VERSION : 0.1
   VAR_INPUT
      SetGroup : Bool;
      "Max Seq Time h_real" : Real;
      "Max Seq Time h" : Time;
      "De-Ox Time h_real" : Real;
      "Re-Ox Time h_real" : Real;
      "Sequence Time h" : Time;
      "Setpoint Time h_real" : Real;
      "Setpoint Time h" : Time;
      "Sequence Time m Offset_real" : Real := 13.0;
      "Sequence Time m Offset" : Time;
      "O2 Confirmed Time_real" : Real;
      "O2 Confirmed Time" : Time;
      "O2 De-Ox Setpoint" : Real;
      "Re-Ox Treatment" : Bool;
      Continue : Bool;   // Continue Sequence After Restart
      Boost : Bool;   // Bypass Sequence Timers
      "Alarm Debounce time" : Time := T#30s;
      "Valve Cycle" : Struct
         Enable : Bool := true;
         Period : Time := T#2h;
         Length : Time := T#30s;
      END_STRUCT;
      "RIO 1" : "3T_IP_DATA";
      "RIO 2" : "2T_IP_DATA";
      "RIO 3" : "2T_IP_DATA";
      "RIO 4" : "2T_IP_DATA";
      "RIO 5" : "2T_IP_DATA";
      "RIO 6" : "2T_IP_DATA";
      "RIO 7" : "1T_IP_DATA";
      RUN : Bool;
      "RUN GROUP 1" : Bool;
      "RUN GROUP 2" : Bool;
      "RUN GROUP 3" : Bool;
      "RUN GROUP 4" : Bool;
      "RUN GROUP 5" : Bool;
      "RUN GROUP 6" : Bool;
      "RUN GROUP 7" : Bool;
      "RUN GROUP 8" : Bool;
      "RUN GROUP 9" : Bool;
      "RUN GROUP 10" : Bool;
      "RUN GROUP 11" : Bool;
      "RUN GROUP 12" : Bool;
      "RUN GROUP 13" : Bool;
      "RUN GROUP 14" : Bool;
      "GROUP ACTIV 1" : Bool;
      "GROUP ACTIV 2" : Bool;
      "GROUP ACTIV 3" : Bool;
      "GROUP ACTIV 4" : Bool;
      "GROUP ACTIV 5" : Bool;
      "GROUP ACTIV 6" : Bool;
      "GROUP ACTIV 7" : Bool;
      "GROUP ACTIV 8" : Bool;
      "GROUP ACTIV 9" : Bool;
      "GROUP ACTIV 10" : Bool;
      "GROUP ACTIV 11" : Bool;
      "GROUP ACTIV 12" : Bool;
      "GROUP ACTIV 13" : Bool;
      "GROUP ACTIV 14" : Bool;
      "TANK ACTIV 1" : Bool;
      "TANK ACTIV 2" : Bool;
      "TANK ACTIV 3" : Bool;
      "TANK ACTIV 4" : Bool;
      "TANK ACTIV 5" : Bool;
      "TANK ACTIV 6" : Bool;
      "TANK ACTIV 7" : Bool;
      "TANK ACTIV 8" : Bool;
      "TANK ACTIV 9" : Bool;
      "TANK ACTIV 10" : Bool;
      "TANK ACTIV 11" : Bool;
      "TANK ACTIV 12" : Bool;
      "TANK ACTIV 13" : Bool;
      "TANK ACTIV 14" : Bool;
      "TANK ACTIV 15" : Bool;
      "TANK ACTIV 16" : Bool;
      "TANK ACTIV 17" : Bool;
      "TANK ACTIV 18" : Bool;
      "TANK ACTIV 19" : Bool;
      "TANK ACTIV 20" : Bool;
      "TANK ACTIV 21" : Bool;
      "TANK ACTIV 22" : Bool;
      "TANK ACTIV 23" : Bool;
      "TANK ACTIV 24" : Bool;
   END_VAR
   VAR_OUTPUT
      "RUN TANK 1" : Bool;
      "RUN TANK 2" : Bool;
      "RUN TANK 3" : Bool;
      "RUN TANK 4" : Bool;
      "RUN TANK 5" : Bool;
      "RUN TANK 6" : Bool;
      "RUN TANK 7" : Bool;
      "RUN TANK 8" : Bool;
      "RUN TANK 9" : Bool;
      "RUN TANK 10" : Bool;
      "RUN TANK 11" : Bool;
      "RUN TANK 12" : Bool;
      "RUN TANK 13" : Bool;
      "RUN TANK 14" : Bool;
      "RUN TANK 15" : Bool;
      "RUN TANK 16" : Bool;
      "RUN TANK 17" : Bool;
      "RUN TANK 18" : Bool;
      "RUN TANK 19" : Bool;
      "RUN TANK 20" : Bool;
      "RUN TANK 21" : Bool;
      "RUN TANK 22" : Bool;
      "RUN TANK 23" : Bool;
      "RUN TANK 24" : Bool;
      "GROUP RUN" : Int;
      "GROUP SET" : Int;
      "GROUP of TANK 1" : Int := 1;
      "GROUP of TANK 2" : Int := 1;
      "GROUP of TANK 3" : Int := 1;
      "GROUP of TANK 4" : Int := 1;
      "GROUP of TANK 5" : Int := 1;
      "GROUP of TANK 6" : Int := 1;
      "GROUP of TANK 7" : Int := 1;
      "GROUP of TANK 8" : Int := 2;
      "GROUP of TANK 9" : Int := 2;
      "GROUP of TANK 10" : Int := 2;
      "GROUP of TANK 11" : Int := 2;
      "GROUP of TANK 12" : Int := 2;
      "GROUP of TANK 13" : Int := 2;
      "GROUP of TANK 14" : Int := 2;
      "GROUP of TANK 15" : Int;
      "GROUP of TANK 16" : Int;
      "GROUP of TANK 17" : Int;
      "GROUP of TANK 18" : Int;
      "GROUP of TANK 19" : Int;
      "GROUP of TANK 20" : Int;
      "GROUP of TANK 21" : Int;
      "GROUP of TANK 22" : Int;
      "GROUP of TANK 23" : Int;
      "GROUP of TANK 24" : Int;
      "Time Left Tank" : Struct
         "Time Left Tank 1" : Real;
         "Time Left Tank 2" : Real;
         "Time Left Tank 3" : Real;
         "Time Left Tank 4" : Real;
         "Time Left Tank 5" : Real;
         "Time Left Tank 6" : Real;
         "Time Left Tank 7" : Real;
         "Time Left Tank 8" : Real;
         "Time Left Tank 9" : Real;
         "Time Left Tank 10" : Real;
         "Time Left Tank 11" : Real;
         "Time Left Tank 12" : Real;
         "Time Left Tank 13" : Real;
         "Time Left Tank 14" : Real;
         "Time Left Tank 15" : Real;
         "Time Left Tank 16" : Real;
         "Time Left Tank 17" : Real;
         "Time Left Tank 18" : Real;
         "Time Left Tank 19" : Real;
         "Time Left Tank 20" : Real;
         "Time Left Tank 21" : Real;
         "Time Left Tank 22" : Real;
         "Time Left Tank 23" : Real;
         "Time Left Tank 24" : Real;
         "Time Left d Tank 1" : DInt;
         "Time Left h Tank 1" : DInt;
         "Time Left m Tank 1" : DInt;
         "Time Left d Tank 2" : DInt;
         "Time Left h Tank 2" : DInt;
         "Time Left m Tank 2" : DInt;
         "Time Left d Tank 3" : DInt;
         "Time Left h Tank 3" : DInt;
         "Time Left m Tank 3" : DInt;
         "Time Left d Tank 4" : DInt;
         "Time Left h Tank 4" : DInt;
         "Time Left m Tank 4" : DInt;
         "Time Left d Tank 5" : DInt;
         "Time Left h Tank 5" : DInt;
         "Time Left m Tank 5" : DInt;
         "Time Left d Tank 6" : DInt;
         "Time Left h Tank 6" : DInt;
         "Time Left m Tank 6" : DInt;
         "Time Left d Tank 7" : DInt;
         "Time Left h Tank 7" : DInt;
         "Time Left m Tank 7" : DInt;
         "Time Left d Tank 8" : DInt;
         "Time Left h Tank 8" : DInt;
         "Time Left m Tank 8" : DInt;
         "Time Left d Tank 9" : DInt;
         "Time Left h Tank 9" : DInt;
         "Time Left m Tank 9" : DInt;
         "Time Left d Tank 10" : DInt;
         "Time Left h Tank 10" : DInt;
         "Time Left m Tank 10" : DInt;
         "Time Left d Tank 11" : DInt;
         "Time Left h Tank 11" : DInt;
         "Time Left m Tank 11" : DInt;
         "Time Left d Tank 12" : DInt;
         "Time Left h Tank 12" : DInt;
         "Time Left m Tank 12" : DInt;
         "Time Left d Tank 13" : DInt;
         "Time Left h Tank 13" : DInt;
         "Time Left m Tank 13" : DInt;
         "Time Left d Tank 14" : DInt;
         "Time Left h Tank 14" : DInt;
         "Time Left m Tank 14" : DInt;
      END_STRUCT;
      "Diff Time Remain" : DInt;
      "GROUP Sequence Done" : Bool;
      "GTT Valves Closed" : Bool;
      "Treatment Time Extend_Hrs" : Time;
      "De-Ox Time Extend_Hrs Real" : Real;
      "Re-Ox Time Extend_Hrs" : Time := T#0ms;
      "Re-Ox Time Extend_Hrs Real" : Real := 0.0;
      "Tank Activ Gr 1" : Bool;
      "Tank Activ Gr 2" : Bool;
      "Tank Activ Gr 3" : Bool;
      "Tank Activ Gr 4" : Bool;
      "Tank Activ Gr 5" : Bool;
      "Tank Activ Gr 6" : Bool;
      "Tank Activ Gr 7" : Bool;
      "Tank Activ Gr 8" : Bool;
      "Tank Activ Gr 9" : Bool;
      "Tank Activ Gr 10" : Bool;
      "Tank Activ Gr 11" : Bool;
      "Tank Activ Gr 12" : Bool;
      "Tank Activ Gr 13" : Bool;
      "Tank Activ Gr 14" : Bool;
      "Tank Activ" : Bool;
   END_VAR
   VAR
      True : Bool;
      False : Bool;
      SetGroupSR : Bool;
      SetGroupFlag : Bool;
      SetGroupDelay : TON_TIME;
      "SET GROUP 1" : Bool;
      "SET GROUP 2" : Bool;
      "SET GROUP 3" : Bool;
      "SET GROUP 4" : Bool;
      "SET GROUP 5" : Bool;
      "SET GROUP 6" : Bool;
      "SET GROUP 7" : Bool;
      "SET GROUP 8" : Bool;
      "SET GROUP 9" : Bool;
      "SET GROUP 10" : Bool;
      "SET GROUP 11" : Bool;
      "SET GROUP 12" : Bool;
      "SET GROUP 13" : Bool;
      "SET GROUP 14" : Bool;
   END_VAR
   VAR RETAIN
      "M GROUP of TANK 1" : Int;
      "M GROUP of TANK 2" : Int;
      "M GROUP of TANK 3" : Int;
      "M GROUP of TANK 4" : Int;
      "M GROUP of TANK 5" : Int;
      "M GROUP of TANK 6" : Int;
      "M GROUP of TANK 7" : Int;
      "M GROUP of TANK 8" : Int;
      "M GROUP of TANK 9" : Int;
      "M GROUP of TANK 10" : Int;
      "M GROUP of TANK 11" : Int;
      "M GROUP of TANK 12" : Int;
      "M GROUP of TANK 13" : Int;
      "M GROUP of TANK 14" : Int;
      "M GROUP of TANK 15" : Int;
      "M GROUP of TANK 16" : Int;
      "M GROUP of TANK 17" : Int;
      "M GROUP of TANK 18" : Int;
      "M GROUP of TANK 19" : Int;
      "M GROUP of TANK 20" : Int;
      "M GROUP of TANK 21" : Int;
      "M GROUP of TANK 22" : Int;
      "M GROUP of TANK 23" : Int;
      "M GROUP of TANK 24" : Int;
   END_VAR
   VAR
      GroupNActivFwdAux : Bool;
      "Change Group Flag" : Bool;
      PulsAuxP : Struct
         "PulsAuxP 1" : Bool;
         "PulsAuxP 2" : Bool;
         "PulsAuxP 3" : Bool;
         "PulsAuxP 4" : Bool;
         "PulsAuxP 5" : Bool;
         "PulsAuxP 6" : Bool;
         "PulsAuxP 7" : Bool;
         "PulsAuxP 8" : Bool;
         "PulsAuxP 9" : Bool;
         "PulsAuxP 10" : Bool;
         "PulsAuxP 11" : Bool;
         "PulsAuxP 12" : Bool;
         "PulsAuxP 13" : Bool;
         "PulsAuxP 14" : Bool;
         "PulsAuxP 15" : Bool;
         "PulsAuxP 16" : Bool;
         "PulsAuxP 17" : Bool;
         "PulsAuxP 18" : Bool;
         "PulsAuxP 19" : Bool;
         "PulsAuxP 20" : Bool;
         "PulsAuxP 21" : Bool;
         "PulsAuxP 22" : Bool;
         "PulsAuxP 23" : Bool;
         "PulsAuxP 24" : Bool;
      END_STRUCT;
      PulsAuxN : Struct
         "PulsAuxN 1" : Bool;
         "PulsAuxN 2" : Bool;
         "PulsAuxN 3" : Bool;
         "PulsAuxN 4" : Bool;
         "PulsAuxN 5" : Bool;
         "PulsAuxN 6" : Bool;
         "PulsAuxN 7" : Bool;
         "PulsAuxN 8" : Bool;
         "PulsAuxN 9" : Bool;
         "PulsAuxN 10" : Bool;
         "PulsAuxN 11" : Bool;
         "PulsAuxN 12" : Bool;
         "PulsAuxN 13" : Bool;
         "PulsAuxN 14" : Bool;
         "PulsAuxN 15" : Bool;
         "PulsAuxN 16" : Bool;
         "PulsAuxN 17" : Bool;
         "PulsAuxN 18" : Bool;
         "PulsAuxN 19" : Bool;
         "PulsAuxN 20" : Bool;
         "PulsAuxN 21" : Bool;
         "PulsAuxN 22" : Bool;
         "PulsAuxN 23" : Bool;
         "PulsAuxN 24" : Bool;
      END_STRUCT;
      "Cycle Tank" : Int;
      "Aux Min Time Tank1" : Bool;
      "Aux Min Time Tank2" : Bool;
      "Aux Min Time Tank3" : Bool;
      "Aux Min Time Tank4" : Bool;
      "Aux Min Time Tank5" : Bool;
      "Aux Min Time Tank6" : Bool;
      "Aux Min Time Tank7" : Bool;
      "Aux Min Time Tank8" : Bool;
      "Aux Min Time Tank9" : Bool;
      "Aux Min Time Tank10" : Bool;
      "Aux Min Time Tank11" : Bool;
      "Aux Min Time Tank12" : Bool;
      "Aux Min Time Tank13" : Bool;
      "Aux Min Time Tank14" : Bool;
      "Aux Min Time Tank15" : Bool;
      "Aux Min Time Tank16" : Bool;
      "Aux Min Time Tank17" : Bool;
      "Aux Min Time Tank18" : Bool;
      "Aux Min Time Tank19" : Bool;
      "Aux Min Time Tank20" : Bool;
      "Aux Min Time Tank21" : Bool;
      "Aux Min Time Tank22" : Bool;
      "Aux Min Time Tank23" : Bool;
      "Aux Min Time Tank24" : Bool;
   END_VAR
   VAR RETAIN
      "GROUP ACTIVE INT 1" : Bool := true;
      "GROUP ACTIVE INT 2" : Bool := true;
      "GROUP ACTIVE INT 3" : Bool := false;
      "GROUP ACTIVE INT 4" : Bool := false;
      "GROUP ACTIVE INT 5" : Bool := false;
      "GROUP ACTIVE INT 6" : Bool := false;
      "GROUP ACTIVE INT 7" : Bool := false;
      "GROUP ACTIVE INT 8" : Bool := false;
      "GROUP ACTIVE INT 9" : Bool := false;
      "GROUP ACTIVE INT 10" : Bool := false;
      "GROUP ACTIVE INT 11" : Bool := false;
      "GROUP ACTIVE INT 12" : Bool := false;
      "GROUP ACTIVE INT 13" : Bool := false;
      "GROUP ACTIVE INT 14" : Bool := false;
   END_VAR
   VAR
      "Sequence Time Min_Aux" : Real;
      "Setpoint Time Min_Aux" : Real;
      "Sequence Time Min Offset_Aux" : Real;
      "O2 Confirmed Time_Aux" : Real;
      "Grup Count" : Int;
      "De-Ox Time Extend_Aux 1" : Real;
      "Max Seq Time h_Aux" : Real;
      "Group Active Flag" : Bool;
      GroupNActivFwd : Bool;
      "Offset Correction Aux" : Real;
   END_VAR
   VAR RETAIN
      "Sequence Time Min Aux" : Struct
         "Sequence Time Min Aux 1" : Time;
         "Sequence Time Min Aux 2" : Time;
         "Sequence Time Min Aux 3" : Time;
         "Sequence Time Min Aux 4" : Time;
         "Sequence Time Min Aux 5" : Time;
         "Sequence Time Min Aux 6" : Time;
         "Sequence Time Min Aux 7" : Time;
         "Sequence Time Min Aux 8" : Time;
         "Sequence Time Min Aux 9" : Time;
         "Sequence Time Min Aux 10" : Time;
         "Sequence Time Min Aux 11" : Time;
         "Sequence Time Min Aux 12" : Time;
         "Sequence Time Min Aux 13" : Time;
         "Sequence Time Min Aux 14" : Time;
         "Sequence Time Min Aux 15" : Time;
         "Sequence Time Min Aux 16" : Time;
         "Sequence Time Min Aux 17" : Time;
         "Sequence Time Min Aux 18" : Time;
         "Sequence Time Min Aux 19" : Time;
         "Sequence Time Min Aux 20" : Time;
         "Sequence Time Min Aux 21" : Time;
         "Sequence Time Min Aux 22" : Time;
         "Sequence Time Min Aux 23" : Time;
         "Sequence Time Min Aux 24" : Time;
      END_STRUCT;
      "Sequence Time Min Memo" : Struct
         "Sequence Time Min Memo 1" : Time;
         "Sequence Time Min Memo 2" : Time;
         "Sequence Time Min Memo 3" : Time;
         "Sequence Time Min Memo 4" : Time;
         "Sequence Time Min Memo 5" : Time;
         "Sequence Time Min Memo 6" : Time;
         "Sequence Time Min Memo 7" : Time;
         "Sequence Time Min Memo 8" : Time;
         "Sequence Time Min Memo 9" : Time;
         "Sequence Time Min Memo 10" : Time;
         "Sequence Time Min Memo 11" : Time;
         "Sequence Time Min Memo 12" : Time;
         "Sequence Time Min Memo 13" : Time;
         "Sequence Time Min Memo 14" : Time;
         "Sequence Time Min Memo 15" : Time;
         "Sequence Time Min Memo 16" : Time;
         "Sequence Time Min Memo 17" : Time;
         "Sequence Time Min Memo 18" : Time;
         "Sequence Time Min Memo 19" : Time;
         "Sequence Time Min Memo 20" : Time;
         "Sequence Time Min Memo 21" : Time;
         "Sequence Time Min Memo 22" : Time;
         "Sequence Time Min Memo 23" : Time;
         "Sequence Time Min Memo 24" : Time;
      END_STRUCT;
   END_VAR
   VAR
      "RUN GROUP ST 1" : Struct
         "RUN TANK 1" : Bool;
         "RUN TANK 2" : Bool;
         "RUN TANK 3" : Bool;
         "RUN TANK 4" : Bool;
         "RUN TANK 5" : Bool;
         "RUN TANK 6" : Bool;
         "RUN TANK 7" : Bool;
         "RUN TANK 8" : Bool;
         "RUN TANK 9" : Bool;
         "RUN TANK 10" : Bool;
         "RUN TANK 11" : Bool;
         "RUN TANK 12" : Bool;
         "RUN TANK 13" : Bool;
         "RUN TANK 14" : Bool;
         "RUN TANK 15" : Bool;
         "RUN TANK 16" : Bool;
         "RUN TANK 17" : Bool;
         "RUN TANK 18" : Bool;
         "RUN TANK 19" : Bool;
         "RUN TANK 20" : Bool;
         "RUN TANK 21" : Bool;
         "RUN TANK 22" : Bool;
         "RUN TANK 23" : Bool;
         "RUN TANK 24" : Bool;
      END_STRUCT;
      "RUN GROUP ST 2" : Struct
         "RUN TANK 1" : Bool;
         "RUN TANK 2" : Bool;
         "RUN TANK 3" : Bool;
         "RUN TANK 4" : Bool;
         "RUN TANK 5" : Bool;
         "RUN TANK 6" : Bool;
         "RUN TANK 7" : Bool;
         "RUN TANK 8" : Bool;
         "RUN TANK 9" : Bool;
         "RUN TANK 10" : Bool;
         "RUN TANK 11" : Bool;
         "RUN TANK 12" : Bool;
         "RUN TANK 13" : Bool;
         "RUN TANK 14" : Bool;
         "RUN TANK 15" : Bool;
         "RUN TANK 16" : Bool;
         "RUN TANK 17" : Bool;
         "RUN TANK 18" : Bool;
         "RUN TANK 19" : Bool;
         "RUN TANK 20" : Bool;
         "RUN TANK 21" : Bool;
         "RUN TANK 22" : Bool;
         "RUN TANK 23" : Bool;
         "RUN TANK 24" : Bool;
      END_STRUCT;
      "RUN GROUP ST 3" : Struct
         "RUN TANK 1" : Bool;
         "RUN TANK 2" : Bool;
         "RUN TANK 3" : Bool;
         "RUN TANK 4" : Bool;
         "RUN TANK 5" : Bool;
         "RUN TANK 6" : Bool;
         "RUN TANK 7" : Bool;
         "RUN TANK 8" : Bool;
         "RUN TANK 9" : Bool;
         "RUN TANK 10" : Bool;
         "RUN TANK 11" : Bool;
         "RUN TANK 12" : Bool;
         "RUN TANK 13" : Bool;
         "RUN TANK 14" : Bool;
         "RUN TANK 15" : Bool;
         "RUN TANK 16" : Bool;
         "RUN TANK 17" : Bool;
         "RUN TANK 18" : Bool;
         "RUN TANK 19" : Bool;
         "RUN TANK 20" : Bool;
         "RUN TANK 21" : Bool;
         "RUN TANK 22" : Bool;
         "RUN TANK 23" : Bool;
         "RUN TANK 24" : Bool;
      END_STRUCT;
      "RUN GROUP ST 4" : Struct
         "RUN TANK 1" : Bool;
         "RUN TANK 2" : Bool;
         "RUN TANK 3" : Bool;
         "RUN TANK 4" : Bool;
         "RUN TANK 5" : Bool;
         "RUN TANK 6" : Bool;
         "RUN TANK 7" : Bool;
         "RUN TANK 8" : Bool;
         "RUN TANK 9" : Bool;
         "RUN TANK 10" : Bool;
         "RUN TANK 11" : Bool;
         "RUN TANK 12" : Bool;
         "RUN TANK 13" : Bool;
         "RUN TANK 14" : Bool;
         "RUN TANK 15" : Bool;
         "RUN TANK 16" : Bool;
         "RUN TANK 17" : Bool;
         "RUN TANK 18" : Bool;
         "RUN TANK 19" : Bool;
         "RUN TANK 20" : Bool;
         "RUN TANK 21" : Bool;
         "RUN TANK 22" : Bool;
         "RUN TANK 23" : Bool;
         "RUN TANK 24" : Bool;
      END_STRUCT;
      "RUN GROUP ST 5" : Struct
         "RUN TANK 1" : Bool;
         "RUN TANK 2" : Bool;
         "RUN TANK 3" : Bool;
         "RUN TANK 4" : Bool;
         "RUN TANK 5" : Bool;
         "RUN TANK 6" : Bool;
         "RUN TANK 7" : Bool;
         "RUN TANK 8" : Bool;
         "RUN TANK 9" : Bool;
         "RUN TANK 10" : Bool;
         "RUN TANK 11" : Bool;
         "RUN TANK 12" : Bool;
         "RUN TANK 13" : Bool;
         "RUN TANK 14" : Bool;
         "RUN TANK 15" : Bool;
         "RUN TANK 16" : Bool;
         "RUN TANK 17" : Bool;
         "RUN TANK 18" : Bool;
         "RUN TANK 19" : Bool;
         "RUN TANK 20" : Bool;
         "RUN TANK 21" : Bool;
         "RUN TANK 22" : Bool;
         "RUN TANK 23" : Bool;
         "RUN TANK 24" : Bool;
      END_STRUCT;
      "RUN GROUP ST 6" : Struct
         "RUN TANK 1" : Bool;
         "RUN TANK 2" : Bool;
         "RUN TANK 3" : Bool;
         "RUN TANK 4" : Bool;
         "RUN TANK 5" : Bool;
         "RUN TANK 6" : Bool;
         "RUN TANK 7" : Bool;
         "RUN TANK 8" : Bool;
         "RUN TANK 9" : Bool;
         "RUN TANK 10" : Bool;
         "RUN TANK 11" : Bool;
         "RUN TANK 12" : Bool;
         "RUN TANK 13" : Bool;
         "RUN TANK 14" : Bool;
         "RUN TANK 15" : Bool;
         "RUN TANK 16" : Bool;
         "RUN TANK 17" : Bool;
         "RUN TANK 18" : Bool;
         "RUN TANK 19" : Bool;
         "RUN TANK 20" : Bool;
         "RUN TANK 21" : Bool;
         "RUN TANK 22" : Bool;
         "RUN TANK 23" : Bool;
         "RUN TANK 24" : Bool;
      END_STRUCT;
      "RUN GROUP ST 7" : Struct
         "RUN TANK 1" : Bool;
         "RUN TANK 2" : Bool;
         "RUN TANK 3" : Bool;
         "RUN TANK 4" : Bool;
         "RUN TANK 5" : Bool;
         "RUN TANK 6" : Bool;
         "RUN TANK 7" : Bool;
         "RUN TANK 8" : Bool;
         "RUN TANK 9" : Bool;
         "RUN TANK 10" : Bool;
         "RUN TANK 11" : Bool;
         "RUN TANK 12" : Bool;
         "RUN TANK 13" : Bool;
         "RUN TANK 14" : Bool;
         "RUN TANK 15" : Bool;
         "RUN TANK 16" : Bool;
         "RUN TANK 17" : Bool;
         "RUN TANK 18" : Bool;
         "RUN TANK 19" : Bool;
         "RUN TANK 20" : Bool;
         "RUN TANK 21" : Bool;
         "RUN TANK 22" : Bool;
         "RUN TANK 23" : Bool;
         "RUN TANK 24" : Bool;
      END_STRUCT;
      "RUN GROUP ST 8" : Struct
         "RUN TANK 1" : Bool;
         "RUN TANK 2" : Bool;
         "RUN TANK 3" : Bool;
         "RUN TANK 4" : Bool;
         "RUN TANK 5" : Bool;
         "RUN TANK 6" : Bool;
         "RUN TANK 7" : Bool;
         "RUN TANK 8" : Bool;
         "RUN TANK 9" : Bool;
         "RUN TANK 10" : Bool;
         "RUN TANK 11" : Bool;
         "RUN TANK 12" : Bool;
         "RUN TANK 13" : Bool;
         "RUN TANK 14" : Bool;
         "RUN TANK 15" : Bool;
         "RUN TANK 16" : Bool;
         "RUN TANK 17" : Bool;
         "RUN TANK 18" : Bool;
         "RUN TANK 19" : Bool;
         "RUN TANK 20" : Bool;
         "RUN TANK 21" : Bool;
         "RUN TANK 22" : Bool;
         "RUN TANK 23" : Bool;
         "RUN TANK 24" : Bool;
      END_STRUCT;
      "RUN GROUP ST 9" : Struct
         "RUN TANK 1" : Bool;
         "RUN TANK 2" : Bool;
         "RUN TANK 3" : Bool;
         "RUN TANK 4" : Bool;
         "RUN TANK 5" : Bool;
         "RUN TANK 6" : Bool;
         "RUN TANK 7" : Bool;
         "RUN TANK 8" : Bool;
         "RUN TANK 9" : Bool;
         "RUN TANK 10" : Bool;
         "RUN TANK 11" : Bool;
         "RUN TANK 12" : Bool;
         "RUN TANK 13" : Bool;
         "RUN TANK 14" : Bool;
         "RUN TANK 15" : Bool;
         "RUN TANK 16" : Bool;
         "RUN TANK 17" : Bool;
         "RUN TANK 18" : Bool;
         "RUN TANK 19" : Bool;
         "RUN TANK 20" : Bool;
         "RUN TANK 21" : Bool;
         "RUN TANK 22" : Bool;
         "RUN TANK 23" : Bool;
         "RUN TANK 24" : Bool;
      END_STRUCT;
      "RUN GROUP ST 10" : Struct
         "RUN TANK 1" : Bool;
         "RUN TANK 2" : Bool;
         "RUN TANK 3" : Bool;
         "RUN TANK 4" : Bool;
         "RUN TANK 5" : Bool;
         "RUN TANK 6" : Bool;
         "RUN TANK 7" : Bool;
         "RUN TANK 8" : Bool;
         "RUN TANK 9" : Bool;
         "RUN TANK 10" : Bool;
         "RUN TANK 11" : Bool;
         "RUN TANK 12" : Bool;
         "RUN TANK 13" : Bool;
         "RUN TANK 14" : Bool;
         "RUN TANK 15" : Bool;
         "RUN TANK 16" : Bool;
         "RUN TANK 17" : Bool;
         "RUN TANK 18" : Bool;
         "RUN TANK 19" : Bool;
         "RUN TANK 20" : Bool;
         "RUN TANK 21" : Bool;
         "RUN TANK 22" : Bool;
         "RUN TANK 23" : Bool;
         "RUN TANK 24" : Bool;
      END_STRUCT;
      "RUN GROUP ST 11" : Struct
         "RUN TANK 1" : Bool;
         "RUN TANK 2" : Bool;
         "RUN TANK 3" : Bool;
         "RUN TANK 4" : Bool;
         "RUN TANK 5" : Bool;
         "RUN TANK 6" : Bool;
         "RUN TANK 7" : Bool;
         "RUN TANK 8" : Bool;
         "RUN TANK 9" : Bool;
         "RUN TANK 10" : Bool;
         "RUN TANK 11" : Bool;
         "RUN TANK 12" : Bool;
         "RUN TANK 13" : Bool;
         "RUN TANK 14" : Bool;
         "RUN TANK 15" : Bool;
         "RUN TANK 16" : Bool;
         "RUN TANK 17" : Bool;
         "RUN TANK 18" : Bool;
         "RUN TANK 19" : Bool;
         "RUN TANK 20" : Bool;
         "RUN TANK 21" : Bool;
         "RUN TANK 22" : Bool;
         "RUN TANK 23" : Bool;
         "RUN TANK 24" : Bool;
      END_STRUCT;
      "RUN GROUP ST 12" : Struct
         "RUN TANK 1" : Bool;
         "RUN TANK 2" : Bool;
         "RUN TANK 3" : Bool;
         "RUN TANK 4" : Bool;
         "RUN TANK 5" : Bool;
         "RUN TANK 6" : Bool;
         "RUN TANK 7" : Bool;
         "RUN TANK 8" : Bool;
         "RUN TANK 9" : Bool;
         "RUN TANK 10" : Bool;
         "RUN TANK 11" : Bool;
         "RUN TANK 12" : Bool;
         "RUN TANK 13" : Bool;
         "RUN TANK 14" : Bool;
         "RUN TANK 15" : Bool;
         "RUN TANK 16" : Bool;
         "RUN TANK 17" : Bool;
         "RUN TANK 18" : Bool;
         "RUN TANK 19" : Bool;
         "RUN TANK 20" : Bool;
         "RUN TANK 21" : Bool;
         "RUN TANK 22" : Bool;
         "RUN TANK 23" : Bool;
         "RUN TANK 24" : Bool;
      END_STRUCT;
      "RUN GROUP ST 13" : Struct
         "RUN TANK 1" : Bool;
         "RUN TANK 2" : Bool;
         "RUN TANK 3" : Bool;
         "RUN TANK 4" : Bool;
         "RUN TANK 5" : Bool;
         "RUN TANK 6" : Bool;
         "RUN TANK 7" : Bool;
         "RUN TANK 8" : Bool;
         "RUN TANK 9" : Bool;
         "RUN TANK 10" : Bool;
         "RUN TANK 11" : Bool;
         "RUN TANK 12" : Bool;
         "RUN TANK 13" : Bool;
         "RUN TANK 14" : Bool;
         "RUN TANK 15" : Bool;
         "RUN TANK 16" : Bool;
         "RUN TANK 17" : Bool;
         "RUN TANK 18" : Bool;
         "RUN TANK 19" : Bool;
         "RUN TANK 20" : Bool;
         "RUN TANK 21" : Bool;
         "RUN TANK 22" : Bool;
         "RUN TANK 23" : Bool;
         "RUN TANK 24" : Bool;
      END_STRUCT;
      "RUN GROUP ST 14" : Struct
         "RUN TANK 1" : Bool;
         "RUN TANK 2" : Bool;
         "RUN TANK 3" : Bool;
         "RUN TANK 4" : Bool;
         "RUN TANK 5" : Bool;
         "RUN TANK 6" : Bool;
         "RUN TANK 7" : Bool;
         "RUN TANK 8" : Bool;
         "RUN TANK 9" : Bool;
         "RUN TANK 10" : Bool;
         "RUN TANK 11" : Bool;
         "RUN TANK 12" : Bool;
         "RUN TANK 13" : Bool;
         "RUN TANK 14" : Bool;
         "RUN TANK 15" : Bool;
         "RUN TANK 16" : Bool;
         "RUN TANK 17" : Bool;
         "RUN TANK 18" : Bool;
         "RUN TANK 19" : Bool;
         "RUN TANK 20" : Bool;
         "RUN TANK 21" : Bool;
         "RUN TANK 22" : Bool;
         "RUN TANK 23" : Bool;
         "RUN TANK 24" : Bool;
      END_STRUCT;
      "Tank1 SP delay" : TOF_TIME;
      "Tank1 Min Time" : TON_TIME;
      "Second Puls" : TP_TIME;
   END_VAR
   VAR RETAIN
      "Group Counter" : CTU_INT;
   END_VAR
   VAR
      "Tank2 Min Time" : TON_TIME;
      "Tank2 SP delay" : TOF_TIME;
      "Tank3 Min Time" : TON_TIME;
      "Tank3 SP delay" : TOF_TIME;
      "Tank4 Min Time" : TON_TIME;
      "Tank4 SP delay" : TOF_TIME;
      "Tank5 Min Time" : TON_TIME;
      "Tank5 SP delay" : TOF_TIME;
      "Tank6 Min Time" : TON_TIME;
      "Tank6 SP delay" : TOF_TIME;
      "Tank7 Min Time" : TON_TIME;
      "Tank7 SP delay" : TOF_TIME;
      "Tank8 Min Time" : TON_TIME;
      "Tank8 SP delay" : TOF_TIME;
      "Tank9 Min Time" : TON_TIME;
      "Tank9 SP delay" : TOF_TIME;
      "Tank10 Min Time" : TON_TIME;
      "Tank10 SP delay" : TOF_TIME;
      "Tank11 Min Time" : TON_TIME;
      "Tank11 SP delay" : TOF_TIME;
      "Tank12 Min Time" : TON_TIME;
      "Tank12 SP delay" : TOF_TIME;
      "Tank13 Min Time" : TON_TIME;
      "Tank13 SP delay" : TOF_TIME;
      "Tank14 Min Time" : TON_TIME;
      "Tank14 SP delay" : TOF_TIME;
      "Tank15 Min Time" : TON_TIME;
      "Tank15 SP delay" : TOF_TIME;
      "Tank16 Min Time" : TON_TIME;
      "Tank16 SP delay" : TOF_TIME;
      "Tank1 O2 Confirm" : TOF_TIME;
      "Tank2 O2 Confirm" : TOF_TIME;
      "Tank3 O2 Confirm" : TOF_TIME;
      "Tank4 O2 Confirm" : TOF_TIME;
      "Tank5 O2 Confirm" : TOF_TIME;
      "Tank6 O2 Confirm" : TOF_TIME;
      "Tank7 O2 Confirm" : TOF_TIME;
      "Tank8 O2 Confirm" : TOF_TIME;
      "Tank9 O2 Confirm" : TOF_TIME;
      "Tank10 O2 Confirm" : TOF_TIME;
      "Tank11 O2 Confirm" : TOF_TIME;
      "Tank12 O2 Confirm" : TOF_TIME;
      "Tank14 O2 Confirm" : TOF_TIME;
      "Tank15 O2 Confirm" : TOF_TIME;
      "Tank16 O2 Confirm" : TOF_TIME;
      "Offset Timer" : TON_TIME;
      "Binary Imputs ADD_Instance" : "Binary Imputs ADD";
      "Activ Groups Number" : "Binary Imputs ADD";
      "Group ActiveFlag" : TON_TIME;
      "Second Puls Timer" : TON_TIME;
      "Sequence Done" : TON_TIME;
      "Tank13 O2 Confirm" : TOF_TIME;
      Choose_Instance_2 : "Choose";
      Choose_Instance_1 : "Choose";
      Choose_Instance_3 : "Choose";
      Choose_Instance_4 : "Choose";
      Choose_Instance_5 : "Choose";
      Choose_Instance_6 : "Choose";
      Choose_Instance_7 : "Choose";
      Choose_Instance_8 : "Choose";
      Choose_Instance_9 : "Choose";
      Choose_Instance_10 : "Choose";
      Choose_Instance_11 : "Choose";
      Choose_Instance_12 : "Choose";
      Choose_Instance_13 : "Choose";
      Choose_Instance_14 : "Choose";
      "Tank1 SP delay II" : TOF_TIME;
      "Tank2 SP delay II" : TOF_TIME;
      "Tank3 SP delay II" : TOF_TIME;
      "Tank4 SP delay II" : TOF_TIME;
      "Tank5 SP delay II" : TOF_TIME;
      "Tank6 SP delay II" : TOF_TIME;
      "Tank7 SP delay II" : TOF_TIME;
      "Tank8 SP delay II" : TOF_TIME;
      "Tank9 SP delay II" : TOF_TIME;
      "Tank10 SP delay II" : TOF_TIME;
      "Tank11 SP delay II" : TOF_TIME;
      "Tank12 SP delay II" : TOF_TIME;
      "Tank13 SP delay II" : TOF_TIME;
      "Tank14 SP delay II" : TOF_TIME;
      "Alarm Tank 1" : TOF_TIME;
      "Alarm Tank 2" : TOF_TIME;
      "Alarm Tank 3" : TOF_TIME;
      "Alarm Tank 4" : TOF_TIME;
      "Alarm Tank 5" : TOF_TIME;
      "Alarm Tank 6" : TOF_TIME;
      "Alarm Tank 7" : TOF_TIME;
      "Alarm Tank 8" : TOF_TIME;
      "Alarm Tank 9" : TOF_TIME;
      "Alarm Tank 10" : TOF_TIME;
      "Alarm Tank 11" : TOF_TIME;
      "Alarm Tank 12" : TOF_TIME;
      "Alarm Tank 13" : TOF_TIME;
      "Alarm Tank 14" : TOF_TIME;
      "Flip Flop Group 14" : "Flip Flop";
      "Flip Flop_1" : "Flip Flop";
      "Flip Flop_2" : "Flip Flop";
      "Flip Flop_3" : "Flip Flop";
      "Flip Flop_4" : "Flip Flop";
      "Flip Flop_5" : "Flip Flop";
      "Flip Flop_6" : "Flip Flop";
      "Flip Flop_7" : "Flip Flop";
      "Flip Flop_8" : "Flip Flop";
      "Flip Flop_9" : "Flip Flop";
      "Flip Flop_10" : "Flip Flop";
      "Flip Flop_11" : "Flip Flop";
      "Flip Flop_12" : "Flip Flop";
      "Flip Flop_13" : "Flip Flop";
      "Flip Flop_14" : "Flip Flop";
      "Flip Flop_15" : "Flip Flop";
      "Flip Flop_16" : "Flip Flop";
      "Flip Flop_17" : "Flip Flop";
      "Flip Flop_18" : "Flip Flop";
      "Flip Flop_19" : "Flip Flop";
      "Flip Flop_20" : "Flip Flop";
      "Flip Flop_21" : "Flip Flop";
      "Flip Flop_22" : "Flip Flop";
      "Flip Flop_23" : "Flip Flop";
      "Flip Flop_24" : "Flip Flop";
      Memory_1 : "Memory";
      Memory_2 : "Memory";
      Memory_3 : "Memory";
      Memory_4 : "Memory";
      Memory_5 : "Memory";
      Memory_6 : "Memory";
      Memory_7 : "Memory";
      Memory_8 : "Memory";
      Memory_9 : "Memory";
      Memory_10 : "Memory";
      Memory_11 : "Memory";
      Memory_12 : "Memory";
      Memory_13 : "Memory";
      Memory_14 : "Memory";
      Memory_15 : "Memory";
      Memory_16 : "Memory";
      Memory_17 : "Memory";
      Memory_18 : "Memory";
      Memory_19 : "Memory";
      Memory_20 : "Memory";
      Memory_21 : "Memory";
      Memory_22 : "Memory";
      Memory_23 : "Memory";
      Memory_24 : "Memory";
      "Cycle Period" : TON_TIME;
      "Cycle Length" : TON_TIME;
   END_VAR
   VAR RETAIN
      "Valve Cycler" : CTU_INT;
      "Cycle Tank Aux" : Int;
   END_VAR
   VAR
      "Sequence Done OutS" : TON_TIME;
      "Hours Timer_1" : "Hours Timer";
      "DInt to Real Calcul #Out := (INT_TO_REAL((#IN1 + #IN2 + #IN3) - (#IN4 + #IN5 + #IN6)) / #IN7)_Instance1" : "DInt to Real Calcul #Out := (INT_TO_REAL((#IN1 + #IN2 + #IN3) - (#IN4 + #IN5 + #IN6)) / #IN7)";
      "DInt to Real Calcul #Out := (INT_TO_REAL((#IN1 + #IN2 + #IN3) - (#IN4 + #IN5 + #IN6)) / #IN7)_Instance2" : "DInt to Real Calcul #Out := (INT_TO_REAL((#IN1 + #IN2 + #IN3) - (#IN4 + #IN5 + #IN6)) / #IN7)";
      "Hours Timer_2" : "Hours Timer";
      "DInt to Real Calcul #Out := (INT_TO_REAL((#IN1 + #IN2 + #IN3) - (#IN4 + #IN5 + #IN6)) / #IN7)_Instance4" : "DInt to Real Calcul #Out := (INT_TO_REAL((#IN1 + #IN2 + #IN3) - (#IN4 + #IN5 + #IN6)) / #IN7)";
      "Hours Timer_4" : "Hours Timer";
      "Hours Timer_3" : "Hours Timer";
      "DInt to Real Calcul #Out := (INT_TO_REAL((#IN1 + #IN2 + #IN3) - (#IN4 + #IN5 + #IN6)) / #IN7)_Instance3" : "DInt to Real Calcul #Out := (INT_TO_REAL((#IN1 + #IN2 + #IN3) - (#IN4 + #IN5 + #IN6)) / #IN7)";
      "DInt to Real Calcul #Out := (INT_TO_REAL((#IN1 + #IN2 + #IN3) - (#IN4 + #IN5 + #IN6)) / #IN7)_Instance5" : "DInt to Real Calcul #Out := (INT_TO_REAL((#IN1 + #IN2 + #IN3) - (#IN4 + #IN5 + #IN6)) / #IN7)";
      "Hours Timer_5" : "Hours Timer";
      "DInt to Real Calcul #Out := (INT_TO_REAL((#IN1 + #IN2 + #IN3) - (#IN4 + #IN5 + #IN6)) / #IN7)_Instance6" : "DInt to Real Calcul #Out := (INT_TO_REAL((#IN1 + #IN2 + #IN3) - (#IN4 + #IN5 + #IN6)) / #IN7)";
      "Hours Timer_6" : "Hours Timer";
      "DInt to Real Calcul #Out := (INT_TO_REAL((#IN1 + #IN2 + #IN3) - (#IN4 + #IN5 + #IN6)) / #IN7)_Instance7" : "DInt to Real Calcul #Out := (INT_TO_REAL((#IN1 + #IN2 + #IN3) - (#IN4 + #IN5 + #IN6)) / #IN7)";
      "Hours Timer_7" : "Hours Timer";
      "DInt to Real Calcul #Out := (INT_TO_REAL((#IN1 + #IN2 + #IN3) - (#IN4 + #IN5 + #IN6)) / #IN7)_Instance8" : "DInt to Real Calcul #Out := (INT_TO_REAL((#IN1 + #IN2 + #IN3) - (#IN4 + #IN5 + #IN6)) / #IN7)";
      "Hours Timer_8" : "Hours Timer";
      "DInt to Real Calcul #Out := (INT_TO_REAL((#IN1 + #IN2 + #IN3) - (#IN4 + #IN5 + #IN6)) / #IN7)_Instance10" : "DInt to Real Calcul #Out := (INT_TO_REAL((#IN1 + #IN2 + #IN3) - (#IN4 + #IN5 + #IN6)) / #IN7)";
      "Hours Timer_10" : "Hours Timer";
      "DInt to Real Calcul #Out := (INT_TO_REAL((#IN1 + #IN2 + #IN3) - (#IN4 + #IN5 + #IN6)) / #IN7)_Instance9" : "DInt to Real Calcul #Out := (INT_TO_REAL((#IN1 + #IN2 + #IN3) - (#IN4 + #IN5 + #IN6)) / #IN7)";
      "Hours Timer_9" : "Hours Timer";
      "DInt to Real Calcul #Out := (INT_TO_REAL((#IN1 + #IN2 + #IN3) - (#IN4 + #IN5 + #IN6)) / #IN7)_Instance11" : "DInt to Real Calcul #Out := (INT_TO_REAL((#IN1 + #IN2 + #IN3) - (#IN4 + #IN5 + #IN6)) / #IN7)";
      "Hours Timer_11" : "Hours Timer";
      "DInt to Real Calcul #Out := (INT_TO_REAL((#IN1 + #IN2 + #IN3) - (#IN4 + #IN5 + #IN6)) / #IN7)_Instance12" : "DInt to Real Calcul #Out := (INT_TO_REAL((#IN1 + #IN2 + #IN3) - (#IN4 + #IN5 + #IN6)) / #IN7)";
      "Hours Timer_12" : "Hours Timer";
      "DInt to Real Calcul #Out := (INT_TO_REAL((#IN1 + #IN2 + #IN3) - (#IN4 + #IN5 + #IN6)) / #IN7)_Instance13" : "DInt to Real Calcul #Out := (INT_TO_REAL((#IN1 + #IN2 + #IN3) - (#IN4 + #IN5 + #IN6)) / #IN7)";
      "Hours Timer_13" : "Hours Timer";
      "DInt to Real Calcul #Out := (INT_TO_REAL((#IN1 + #IN2 + #IN3) - (#IN4 + #IN5 + #IN6)) / #IN7)_Instance14" : "DInt to Real Calcul #Out := (INT_TO_REAL((#IN1 + #IN2 + #IN3) - (#IN4 + #IN5 + #IN6)) / #IN7)";
      "Hours Timer_14" : "Hours Timer";
   END_VAR
   VAR_TEMP   // added for the SCL form of the ladder/FBD networks
      _w1 : Bool;
      _w2 : Bool;
      _w3 : Bool;
      _w4 : Bool;
      _w5 : Bool;
      _w6 : Bool;
      _w7 : Bool;
      _w8 : Bool;
      _w9 : Bool;
      _w10 : Bool;
      _w11 : Bool;
      _w12 : Bool;
      _w13 : Bool;
      _w14 : Bool;
      _w15 : Bool;
      _w16 : Bool;
      _w17 : Bool;
      _w18 : Bool;
      _w19 : Bool;
      _w20 : Bool;
      _w21 : Bool;
      _w22 : Bool;
      _w23 : Bool;
      _w24 : Bool;
      _w25 : Bool;
      _w26 : Bool;
      _w27 : Bool;
      _w28 : Bool;
      _w29 : Bool;
      _w30 : Bool;
      _w31 : Bool;
      _w32 : Bool;
      _w33 : Bool;
      _w34 : Bool;
      _w35 : Bool;
      _w36 : Bool;
      _w37 : Bool;
      _w38 : Bool;
      _w39 : Bool;
      _w40 : Bool;
      _w41 : Bool;
      _w42 : Bool;
      _w43 : Bool;
      _w44 : Bool;
      _w45 : Bool;
      _w46 : Bool;
      _w47 : Bool;
      _w48 : Bool;
      _w49 : Bool;
      _w50 : Bool;
      _w51 : Bool;
      _w52 : Bool;
      _w53 : Bool;
      _w54 : Bool;
      _w55 : Bool;
      _w56 : Bool;
      _w57 : Bool;
      _w58 : Bool;
      _w59 : Bool;
      _w60 : Bool;
      _w61 : Bool;
      _w62 : Bool;
      _w63 : Bool;
      _w64 : Bool;
      _w65 : Bool;
      _w66 : Bool;
      _w67 : Bool;
      _w68 : Bool;
      _w69 : Bool;
      _w70 : Bool;
      _w71 : Bool;
      _w72 : Bool;
   END_VAR
BEGIN

REGION Network 1: False/True
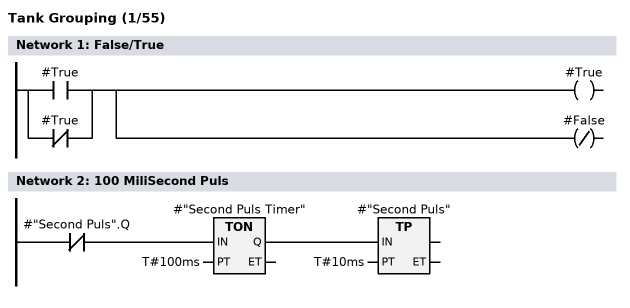
   RUNG wire#powerrail
      Contact( #True )
      wire#w1
      Coil( #True )
   END_RUNG
   RUNG wire#powerrail
      I_Contact( #True )
   END_RUNG wire#w1
   RUNG wire#w1
      I_Coil( #False )
   END_RUNG
   // the same network as SCL:
   #True := #True OR NOT #True;
   #False := NOT #True;
END_REGION

REGION Network 2: 100 MiliSecond Puls
   #"Second Puls Timer"(IN := NOT #"Second Puls".Q, PT := T#100ms);   // TON
   #"Second Puls"(IN := #"Second Puls Timer".Q, PT := T#10ms);   // TP
END_REGION

REGION Network 3: Alarm Debounce
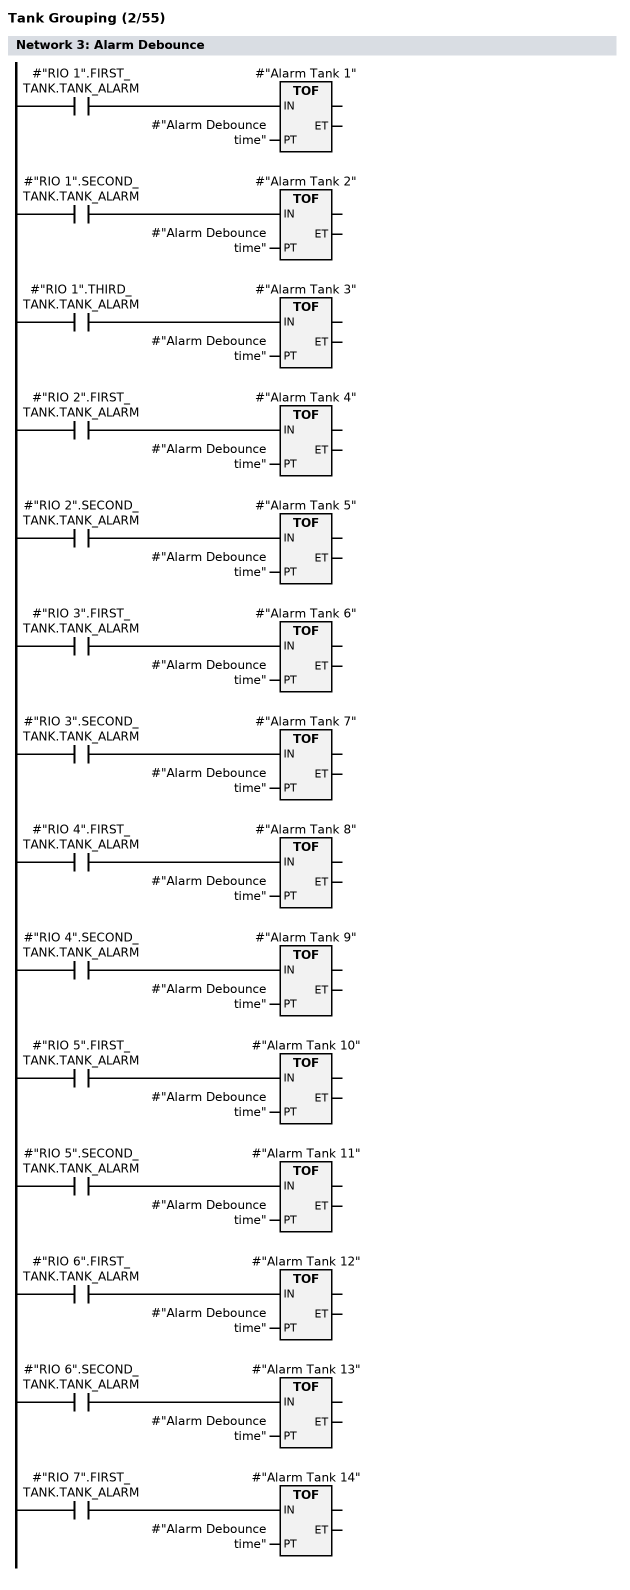
   #"Alarm Tank 1"(IN := #"RIO 1".FIRST_TANK.TANK_ALARM, PT := #"Alarm Debounce time");   // TOF
   #"Alarm Tank 2"(IN := #"RIO 1".SECOND_TANK.TANK_ALARM, PT := #"Alarm Debounce time");   // TOF
   #"Alarm Tank 3"(IN := #"RIO 1".THIRD_TANK.TANK_ALARM, PT := #"Alarm Debounce time");   // TOF
   #"Alarm Tank 4"(IN := #"RIO 2".FIRST_TANK.TANK_ALARM, PT := #"Alarm Debounce time");   // TOF
   #"Alarm Tank 5"(IN := #"RIO 2".SECOND_TANK.TANK_ALARM, PT := #"Alarm Debounce time");   // TOF
   #"Alarm Tank 6"(IN := #"RIO 3".FIRST_TANK.TANK_ALARM, PT := #"Alarm Debounce time");   // TOF
   #"Alarm Tank 7"(IN := #"RIO 3".SECOND_TANK.TANK_ALARM, PT := #"Alarm Debounce time");   // TOF
   #"Alarm Tank 8"(IN := #"RIO 4".FIRST_TANK.TANK_ALARM, PT := #"Alarm Debounce time");   // TOF
   #"Alarm Tank 9"(IN := #"RIO 4".SECOND_TANK.TANK_ALARM, PT := #"Alarm Debounce time");   // TOF
   #"Alarm Tank 10"(IN := #"RIO 5".FIRST_TANK.TANK_ALARM, PT := #"Alarm Debounce time");   // TOF
   #"Alarm Tank 11"(IN := #"RIO 5".SECOND_TANK.TANK_ALARM, PT := #"Alarm Debounce time");   // TOF
   #"Alarm Tank 12"(IN := #"RIO 6".FIRST_TANK.TANK_ALARM, PT := #"Alarm Debounce time");   // TOF
   #"Alarm Tank 13"(IN := #"RIO 6".SECOND_TANK.TANK_ALARM, PT := #"Alarm Debounce time");   // TOF
   #"Alarm Tank 14"(IN := #"RIO 7".FIRST_TANK.TANK_ALARM, PT := #"Alarm Debounce time");   // TOF
END_REGION

REGION Network 4: Set Group SR
   // HMI Button to be set as SetTagWhileKeyPres
